// TIA Portal project "CLU" (V13) (continued)
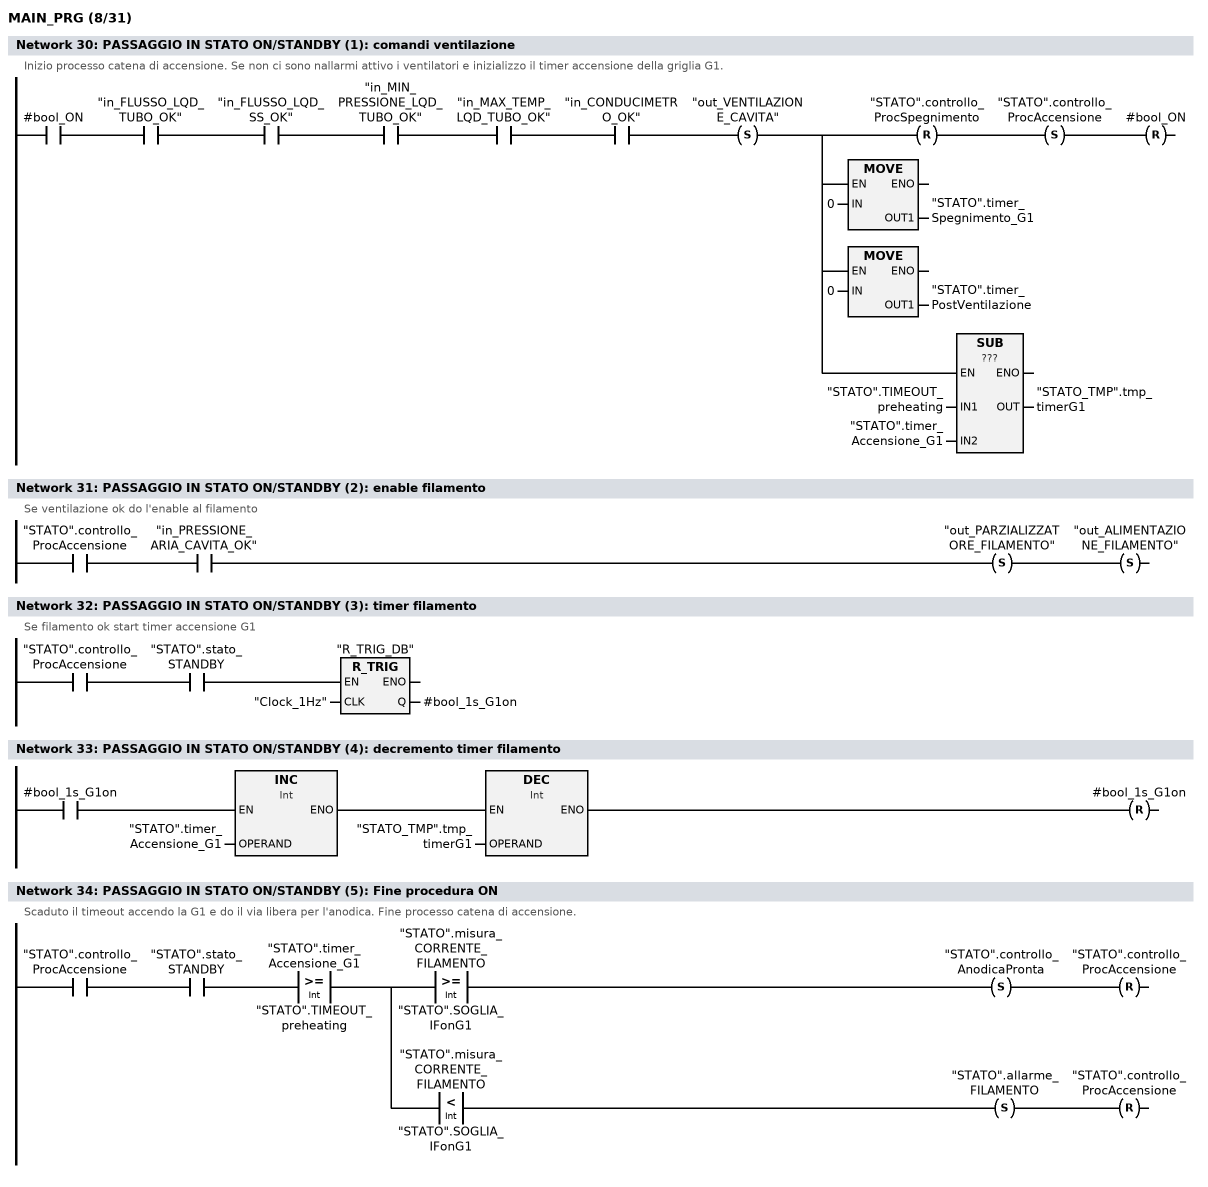
   RUNG wire#powerrail
      Contact( #bool_ON )
      Contact( "in_FLUSSO_LQD_TUBO_OK" )
      Contact( "in_FLUSSO_LQD_SS_OK" )
      Contact( "in_MIN_PRESSIONE_LQD_TUBO_OK" )
      Contact( "in_MAX_TEMP_LQD_TUBO_OK" )
      Contact( "in_CONDUCIMETRO_OK" )
      S_Coil( "out_VENTILAZIONE_CAVITA" )
      wire#w1
      R_Coil( "STATO".controllo_ProcSpegnimento )
      S_Coil( "STATO".controllo_ProcAccensione )
      R_Coil( #bool_ON )
   END_RUNG
   RUNG wire#w1
      Move(in := 0, out1 => "STATO".timer_Spegnimento_G1)
   END_RUNG
   RUNG wire#w1
      Move(in := 0, out1 => "STATO".timer_PostVentilazione)
   END_RUNG
   RUNG wire#w1
      { S7_Templates := "SrcType := ???" } Sub(in1 := "STATO".TIMEOUT_preheating, in2 := "STATO".timer_Accensione_G1, out => "STATO_TMP".tmp_timerG1)
   END_RUNG
   // the same network as SCL:
   IF #bool_ON AND "in_FLUSSO_LQD_TUBO_OK" AND "in_FLUSSO_LQD_SS_OK" AND "in_MIN_PRESSIONE_LQD_TUBO_OK" AND "in_MAX_TEMP_LQD_TUBO_OK" AND "in_CONDUCIMETRO_OK" THEN
       "out_VENTILAZIONE_CAVITA" := TRUE;
       "STATO".controllo_ProcSpegnimento := FALSE;
       "STATO".controllo_ProcAccensione := TRUE;
   END_IF;
   #_w1 := #bool_ON AND "in_FLUSSO_LQD_TUBO_OK" AND "in_FLUSSO_LQD_SS_OK" AND "in_MIN_PRESSIONE_LQD_TUBO_OK" AND "in_MAX_TEMP_LQD_TUBO_OK" AND "in_CONDUCIMETRO_OK";
   IF #_w1 THEN
       #bool_ON := FALSE;
       "STATO".timer_Spegnimento_G1 := 0;
       "STATO".timer_PostVentilazione := 0;
       "STATO_TMP".tmp_timerG1 := "STATO".TIMEOUT_preheating - "STATO".timer_Accensione_G1;
   END_IF;
END_REGION

REGION Network 31: PASSAGGIO IN STATO ON/STANDBY (2): enable filamento
   // Se ventilazione ok do l'enable al filamento
   RUNG wire#powerrail
      Contact( "STATO".controllo_ProcAccensione )
      Contact( "in_PRESSIONE_ARIA_CAVITA_OK" )
      S_Coil( "out_PARZIALIZZATORE_FILAMENTO" )
      S_Coil( "out_ALIMENTAZIONE_FILAMENTO" )
   END_RUNG
   // the same network as SCL:
   IF "STATO".controllo_ProcAccensione AND "in_PRESSIONE_ARIA_CAVITA_OK" THEN
       "out_PARZIALIZZATORE_FILAMENTO" := TRUE;
       "out_ALIMENTAZIONE_FILAMENTO" := TRUE;
   END_IF;
END_REGION

REGION Network 32: PASSAGGIO IN STATO ON/STANDBY (3): timer filamento
   // Se filamento ok start timer accensione G1
   IF "STATO".controllo_ProcAccensione AND "STATO".stato_STANDBY THEN
       "R_TRIG_DB"(CLK := "Clock_1Hz", Q => #bool_1s_G1on);   // R_TRIG
   END_IF;
END_REGION

REGION Network 33: PASSAGGIO IN STATO ON/STANDBY (4): decremento timer filamento
   RUNG wire#powerrail
      Contact( #bool_1s_G1on )
      { S7_Templates := "DestType := Int" } Inc( "STATO".timer_Accensione_G1 )
      { S7_Templates := "DestType := Int" } Dec( "STATO_TMP".tmp_timerG1 )
      R_Coil( #bool_1s_G1on )
   END_RUNG
   // the same network as SCL:
   IF #bool_1s_G1on THEN
       "STATO".timer_Accensione_G1 := "STATO".timer_Accensione_G1 + 1;
       "STATO_TMP".tmp_timerG1 := "STATO_TMP".tmp_timerG1 - 1;
       #bool_1s_G1on := FALSE;
   END_IF;
END_REGION

REGION Network 34: PASSAGGIO IN STATO ON/STANDBY (5): Fine procedura ON
   // Scaduto il timeout accendo la G1 e do il via libera per l'anodica. Fine processo catena di accensione.
   RUNG wire#powerrail
      Contact( "STATO".controllo_ProcAccensione )
      Contact( "STATO".stato_STANDBY )
      { S7_Templates := "SrcType := Int" } GE_Contact(in1 := "STATO".timer_Accensione_G1, in2 := "STATO".TIMEOUT_preheating)
      wire#w1
      { S7_Templates := "SrcType := Int" } GE_Contact(in1 := "STATO".misura_CORRENTE_FILAMENTO, in2 := "STATO".SOGLIA_IFonG1)
      S_Coil( "STATO".controllo_AnodicaPronta )
      R_Coil( "STATO".controllo_ProcAccensione )
   END_RUNG
   RUNG wire#w1
      { S7_Templates := "SrcType := Int" } LT_Contact(in1 := "STATO".misura_CORRENTE_FILAMENTO, in2 := "STATO".SOGLIA_IFonG1)
      S_Coil( "STATO".allarme_FILAMENTO )
      R_Coil( "STATO".controllo_ProcAccensione )
   END_RUNG
   // the same network as SCL:
   #_w1 := "STATO".controllo_ProcAccensione AND "STATO".stato_STANDBY AND ("STATO".timer_Accensione_G1 >= "STATO".TIMEOUT_preheating);
   IF #_w1 AND ("STATO".misura_CORRENTE_FILAMENTO >= "STATO".SOGLIA_IFonG1) THEN
       "STATO".controllo_AnodicaPronta := TRUE;
       "STATO".controllo_ProcAccensione := FALSE;
   END_IF;
   IF #_w1 AND ("STATO".misura_CORRENTE_FILAMENTO < "STATO".SOGLIA_IFonG1) THEN
       "STATO".allarme_FILAMENTO := TRUE;
       "STATO".controllo_ProcAccensione := FALSE;
   END_IF;
END_REGION

REGION Network 35: PASSAGGIO IN ANODICA ON (1): inizio accensione anodica
   // Se il processo catena di accensione è terminato posso iniziare il processo catena di accensione anodica.
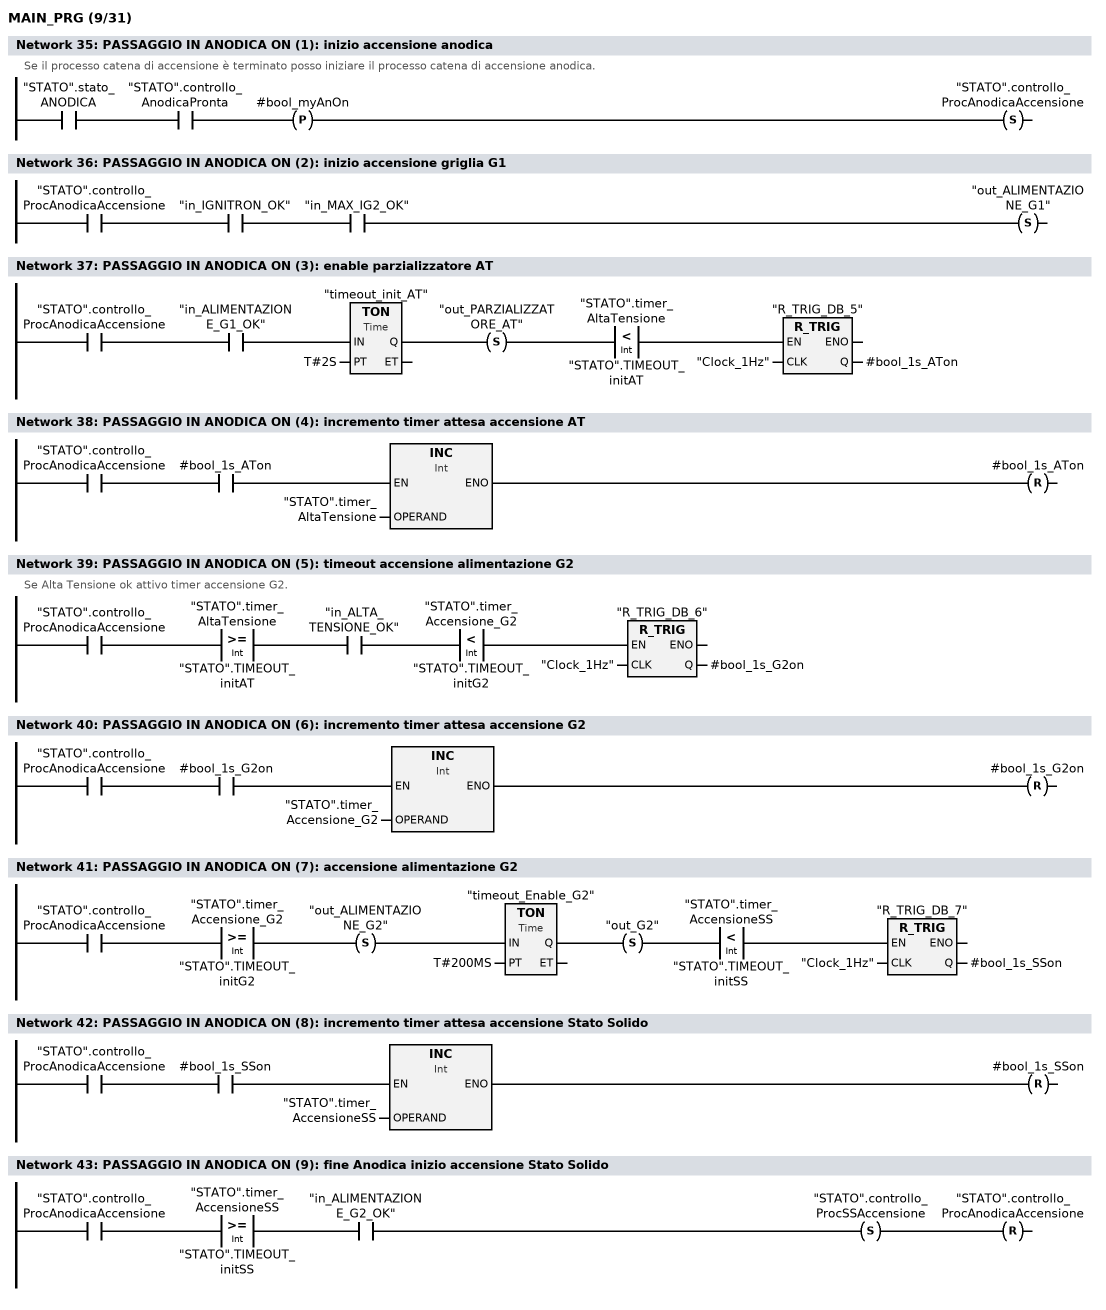
   RUNG wire#powerrail
      Contact( "STATO".stato_ANODICA )
      Contact( "STATO".controllo_AnodicaPronta )
      P_Trig( #bool_myAnOn )
      S_Coil( "STATO".controllo_ProcAnodicaAccensione )
   END_RUNG
   // the same network as SCL:
   #_w1 := "STATO".stato_ANODICA AND "STATO".controllo_AnodicaPronta;
   #_w2 := #_w1 AND NOT #bool_myAnOn;   // rising edge
   #bool_myAnOn := #_w1;
   IF #_w2 THEN "STATO".controllo_ProcAnodicaAccensione := TRUE; END_IF;
END_REGION

REGION Network 36: PASSAGGIO IN ANODICA ON (2): inizio accensione griglia G1
   RUNG wire#powerrail
      Contact( "STATO".controllo_ProcAnodicaAccensione )
      Contact( "in_IGNITRON_OK" )
      Contact( "in_MAX_IG2_OK" )
      S_Coil( "out_ALIMENTAZIONE_G1" )
   END_RUNG
   // the same network as SCL:
   IF "STATO".controllo_ProcAnodicaAccensione AND "in_IGNITRON_OK" AND "in_MAX_IG2_OK" THEN
       "out_ALIMENTAZIONE_G1" := TRUE;
   END_IF;
END_REGION

REGION Network 37: PASSAGGIO IN ANODICA ON (3): enable parzializzatore AT
   "timeout_init_AT".TON(IN := "STATO".controllo_ProcAnodicaAccensione AND "in_ALIMENTAZIONE_G1_OK", PT := T#2S);
   IF "timeout_init_AT".Q THEN "out_PARZIALIZZATORE_AT" := TRUE; END_IF;
   IF "timeout_init_AT".Q AND ("STATO".timer_AltaTensione < "STATO".TIMEOUT_initAT) THEN
       "R_TRIG_DB_5"(CLK := "Clock_1Hz", Q => #bool_1s_ATon);   // R_TRIG
   END_IF;
END_REGION

REGION Network 38: PASSAGGIO IN ANODICA ON (4): incremento timer attesa accensione AT
   RUNG wire#powerrail
      Contact( "STATO".controllo_ProcAnodicaAccensione )
      Contact( #bool_1s_ATon )
      { S7_Templates := "DestType := Int" } Inc( "STATO".timer_AltaTensione )
      R_Coil( #bool_1s_ATon )
   END_RUNG
   // the same network as SCL:
   IF "STATO".controllo_ProcAnodicaAccensione AND #bool_1s_ATon THEN
       "STATO".timer_AltaTensione := "STATO".timer_AltaTensione + 1;
       #bool_1s_ATon := FALSE;
   END_IF;
END_REGION

REGION Network 39: PASSAGGIO IN ANODICA ON (5): timeout accensione alimentazione G2
   // Se Alta Tensione ok attivo timer accensione G2.
   IF "STATO".controllo_ProcAnodicaAccensione AND ("STATO".timer_AltaTensione >= "STATO".TIMEOUT_initAT) AND "in_ALTA_TENSIONE_OK" AND ("STATO".timer_Accensione_G2 < "STATO".TIMEOUT_initG2) THEN
       "R_TRIG_DB_6"(CLK := "Clock_1Hz", Q => #bool_1s_G2on);   // R_TRIG
   END_IF;
END_REGION

REGION Network 40: PASSAGGIO IN ANODICA ON (6): incremento timer attesa accensione G2
   RUNG wire#powerrail
      Contact( "STATO".controllo_ProcAnodicaAccensione )
      Contact( #bool_1s_G2on )
      { S7_Templates := "DestType := Int" } Inc( "STATO".timer_Accensione_G2 )
      R_Coil( #bool_1s_G2on )
   END_RUNG
   // the same network as SCL:
   IF "STATO".controllo_ProcAnodicaAccensione AND #bool_1s_G2on THEN
       "STATO".timer_Accensione_G2 := "STATO".timer_Accensione_G2 + 1;
       #bool_1s_G2on := FALSE;
   END_IF;
END_REGION

REGION Network 41: PASSAGGIO IN ANODICA ON (7): accensione alimentazione G2
   #_w1 := "STATO".controllo_ProcAnodicaAccensione AND ("STATO".timer_Accensione_G2 >= "STATO".TIMEOUT_initG2);
   IF #_w1 THEN "out_ALIMENTAZIONE_G2" := TRUE; END_IF;
   "timeout_Enable_G2".TON(IN := #_w1, PT := T#200MS);
   IF "timeout_Enable_G2".Q THEN "out_G2" := TRUE; END_IF;
   IF "timeout_Enable_G2".Q AND ("STATO".timer_AccensioneSS < "STATO".TIMEOUT_initSS) THEN
       "R_TRIG_DB_7"(CLK := "Clock_1Hz", Q => #bool_1s_SSon);   // R_TRIG
   END_IF;
END_REGION

REGION Network 42: PASSAGGIO IN ANODICA ON (8): incremento timer attesa accensione Stato Solido
   RUNG wire#powerrail
      Contact( "STATO".controllo_ProcAnodicaAccensione )
      Contact( #bool_1s_SSon )
      { S7_Templates := "DestType := Int" } Inc( "STATO".timer_AccensioneSS )
      R_Coil( #bool_1s_SSon )
   END_RUNG
   // the same network as SCL:
   IF "STATO".controllo_ProcAnodicaAccensione AND #bool_1s_SSon THEN
       "STATO".timer_AccensioneSS := "STATO".timer_AccensioneSS + 1;
       #bool_1s_SSon := FALSE;
   END_IF;
END_REGION

REGION Network 43: PASSAGGIO IN ANODICA ON (9): fine Anodica inizio accensione Stato Solido
   RUNG wire#powerrail
      Contact( "STATO".controllo_ProcAnodicaAccensione )
      { S7_Templates := "SrcType := Int" } GE_Contact(in1 := "STATO".timer_AccensioneSS, in2 := "STATO".TIMEOUT_initSS)
      Contact( "in_ALIMENTAZIONE_G2_OK" )
      S_Coil( "STATO".controllo_ProcSSAccensione )
      R_Coil( "STATO".controllo_ProcAnodicaAccensione )
   END_RUNG
   // the same network as SCL:
   IF "STATO".controllo_ProcAnodicaAccensione AND ("STATO".timer_AccensioneSS >= "STATO".TIMEOUT_initSS) AND "in_ALIMENTAZIONE_G2_OK" THEN
       "STATO".controllo_ProcSSAccensione := TRUE;
       "STATO".controllo_ProcAnodicaAccensione := FALSE;
   END_IF;
END_REGION

REGION Network 44: ACCENSIONE STATO SOLIDO (1): accensione amplificatore (impulsivo) AMP 1
   // Se modalità  impulsiva attiva accendo gli amplificatori e attivo timer accensione driver.
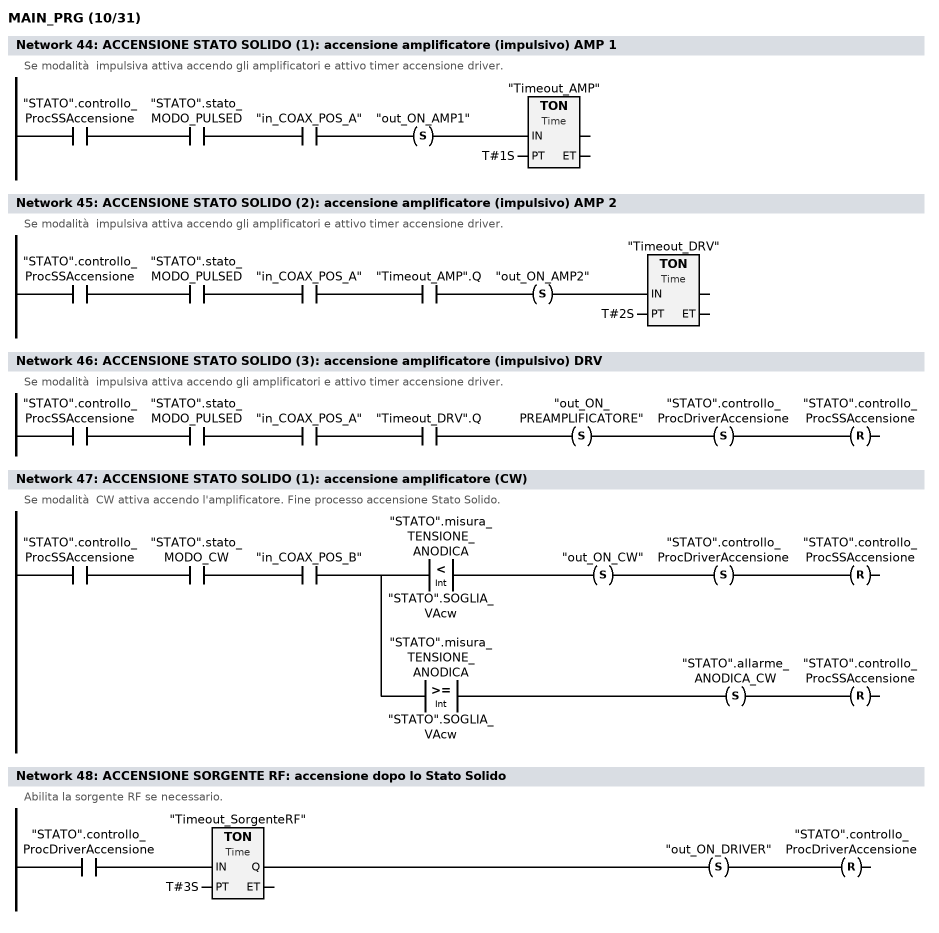
   #_w1 := "STATO".controllo_ProcSSAccensione AND "STATO".stato_MODO_PULSED AND "in_COAX_POS_A";
   IF #_w1 THEN "out_ON_AMP1" := TRUE; END_IF;
   "Timeout_AMP".TON(IN := #_w1, PT := T#1S);
END_REGION

REGION Network 45: ACCENSIONE STATO SOLIDO (2): accensione amplificatore (impulsivo) AMP 2
   // Se modalità  impulsiva attiva accendo gli amplificatori e attivo timer accensione driver.
   #_w1 := "STATO".controllo_ProcSSAccensione AND "STATO".stato_MODO_PULSED AND "in_COAX_POS_A" AND "Timeout_AMP".Q;
   IF #_w1 THEN "out_ON_AMP2" := TRUE; END_IF;
   "Timeout_DRV".TON(IN := #_w1, PT := T#2S);
END_REGION

REGION Network 46: ACCENSIONE STATO SOLIDO (3): accensione amplificatore (impulsivo) DRV
   // Se modalità  impulsiva attiva accendo gli amplificatori e attivo timer accensione driver.
   RUNG wire#powerrail
      Contact( "STATO".controllo_ProcSSAccensione )
      Contact( "STATO".stato_MODO_PULSED )
      Contact( "in_COAX_POS_A" )
      Contact( "Timeout_DRV".Q )
      S_Coil( "out_ON_PREAMPLIFICATORE" )
      S_Coil( "STATO".controllo_ProcDriverAccensione )
      R_Coil( "STATO".controllo_ProcSSAccensione )
   END_RUNG
   // the same network as SCL:
   IF "STATO".controllo_ProcSSAccensione AND "STATO".stato_MODO_PULSED AND "in_COAX_POS_A" AND "Timeout_DRV".Q THEN
       "out_ON_PREAMPLIFICATORE" := TRUE;
       "STATO".controllo_ProcDriverAccensione := TRUE;
       "STATO".controllo_ProcSSAccensione := FALSE;
   END_IF;
END_REGION

REGION Network 47: ACCENSIONE STATO SOLIDO (1): accensione amplificatore (CW)
   // Se modalità  CW attiva accendo l'amplificatore. Fine processo accensione Stato Solido.
   RUNG wire#powerrail
      Contact( "STATO".controllo_ProcSSAccensione )
      Contact( "STATO".stato_MODO_CW )
      Contact( "in_COAX_POS_B" )
      wire#w1
      { S7_Templates := "SrcType := Int" } LT_Contact(in1 := "STATO".misura_TENSIONE_ANODICA, in2 := "STATO".SOGLIA_VAcw)
      S_Coil( "out_ON_CW" )
      S_Coil( "STATO".controllo_ProcDriverAccensione )
      R_Coil( "STATO".controllo_ProcSSAccensione )
   END_RUNG
   RUNG wire#w1
      { S7_Templates := "SrcType := Int" } GE_Contact(in1 := "STATO".misura_TENSIONE_ANODICA, in2 := "STATO".SOGLIA_VAcw)
      S_Coil( "STATO".allarme_ANODICA_CW )
      R_Coil( "STATO".controllo_ProcSSAccensione )
   END_RUNG
   // the same network as SCL:
   #_w1 := "STATO".controllo_ProcSSAccensione AND "STATO".stato_MODO_CW AND "in_COAX_POS_B";
   IF #_w1 AND ("STATO".misura_TENSIONE_ANODICA < "STATO".SOGLIA_VAcw) THEN
       "out_ON_CW" := TRUE;
       "STATO".controllo_ProcDriverAccensione := TRUE;
       "STATO".controllo_ProcSSAccensione := FALSE;
   END_IF;
   IF #_w1 AND ("STATO".misura_TENSIONE_ANODICA >= "STATO".SOGLIA_VAcw) THEN
       "STATO".allarme_ANODICA_CW := TRUE;
       "STATO".controllo_ProcSSAccensione := FALSE;
   END_IF;
END_REGION

REGION Network 48: ACCENSIONE SORGENTE RF: accensione dopo lo Stato Solido
   // Abilita la sorgente RF se necessario.
   "Timeout_SorgenteRF".TON(IN := "STATO".controllo_ProcDriverAccensione, PT := T#3S);
   IF "Timeout_SorgenteRF".Q THEN
       "out_ON_DRIVER" := TRUE;
       "STATO".controllo_ProcDriverAccensione := FALSE;
   END_IF;
END_REGION

REGION Network 49: PASSAGGIO IN ANODICA OFF (1): spegnimento Stato Solido e alimentazione G2
   // Spengo Stato Solido (CW o impulsivo) e alimentazione G2. Inizio processo catena di spegnimento Anodica.
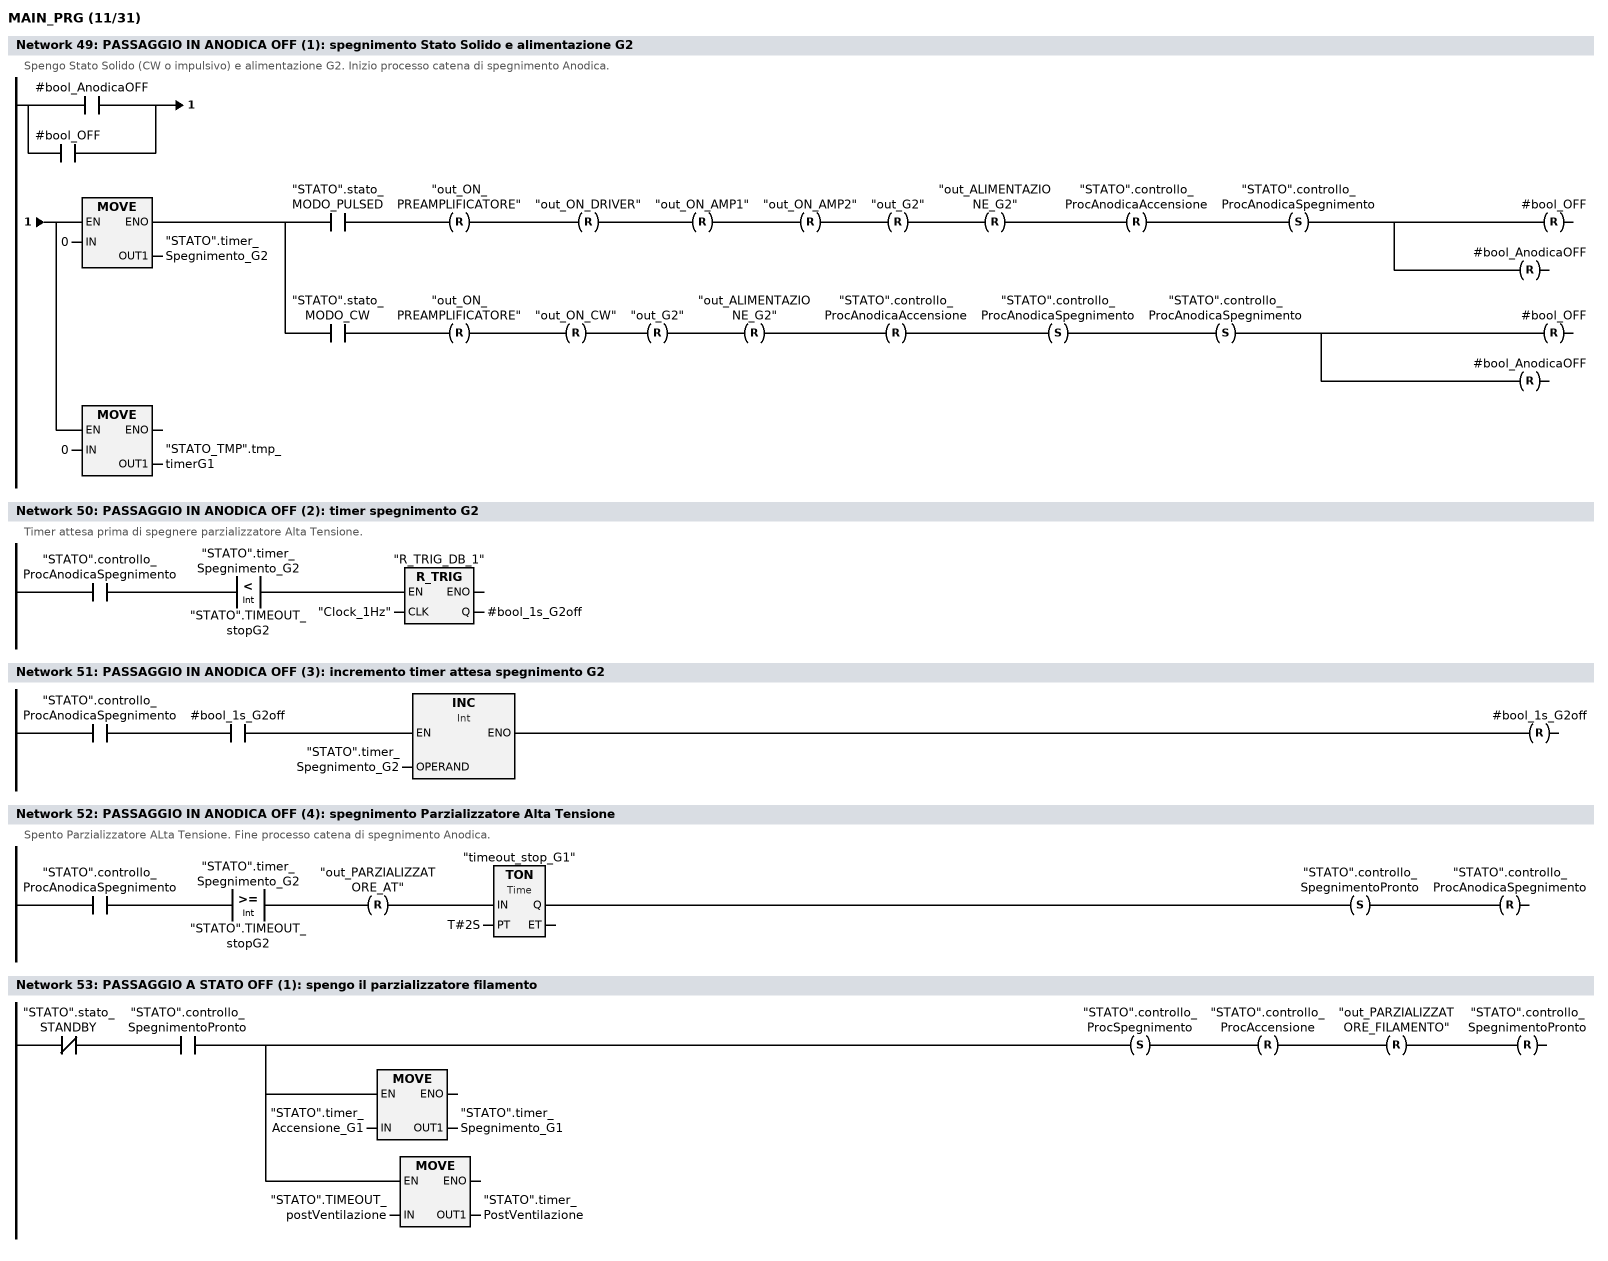
   RUNG wire#powerrail
      Contact( #bool_AnodicaOFF )
      wire#w1
      Move(in := 0, out1 => "STATO".timer_Spegnimento_G2)
      wire#w2
      Contact( "STATO".stato_MODO_PULSED )
      R_Coil( "out_ON_PREAMPLIFICATORE" )
      R_Coil( "out_ON_DRIVER" )
      R_Coil( "out_ON_AMP1" )
      R_Coil( "out_ON_AMP2" )
      R_Coil( "out_G2" )
      R_Coil( "out_ALIMENTAZIONE_G2" )
      R_Coil( "STATO".controllo_ProcAnodicaAccensione )
      S_Coil( "STATO".controllo_ProcAnodicaSpegnimento )
      wire#w3
      R_Coil( #bool_OFF )
   END_RUNG
   RUNG wire#powerrail
      Contact( #bool_OFF )
   END_RUNG wire#w1
   RUNG wire#w3
      R_Coil( #bool_AnodicaOFF )
   END_RUNG
   RUNG wire#w2
      Contact( "STATO".stato_MODO_CW )
      R_Coil( "out_ON_PREAMPLIFICATORE" )
      R_Coil( "out_ON_CW" )
      R_Coil( "out_G2" )
      R_Coil( "out_ALIMENTAZIONE_G2" )
      R_Coil( "STATO".controllo_ProcAnodicaAccensione )
      S_Coil( "STATO".controllo_ProcAnodicaSpegnimento )
      S_Coil( "STATO".controllo_ProcAnodicaSpegnimento )
      wire#w4
      R_Coil( #bool_OFF )
   END_RUNG
   RUNG wire#w4
      R_Coil( #bool_AnodicaOFF )
   END_RUNG
   RUNG wire#w1
      Move(in := 0, out1 => "STATO_TMP".tmp_timerG1)
   END_RUNG
   // the same network as SCL:
   #_w1 := #bool_AnodicaOFF OR #bool_OFF;
   IF #_w1 THEN "STATO".timer_Spegnimento_G2 := 0; END_IF;
   IF #_w1 AND "STATO".stato_MODO_PULSED THEN
       "out_ON_PREAMPLIFICATORE" := FALSE;
       "out_ON_DRIVER" := FALSE;
       "out_ON_AMP1" := FALSE;
       "out_ON_AMP2" := FALSE;
       "out_G2" := FALSE;
       "out_ALIMENTAZIONE_G2" := FALSE;
       "STATO".controllo_ProcAnodicaAccensione := FALSE;
       "STATO".controllo_ProcAnodicaSpegnimento := TRUE;
       #bool_OFF := FALSE;
       #bool_AnodicaOFF := FALSE;
   END_IF;
   IF #_w1 AND "STATO".stato_MODO_CW THEN
       "out_ON_PREAMPLIFICATORE" := FALSE;
       "out_ON_CW" := FALSE;
       "out_G2" := FALSE;
       "out_ALIMENTAZIONE_G2" := FALSE;
       "STATO".controllo_ProcAnodicaAccensione := FALSE;
       "STATO".controllo_ProcAnodicaSpegnimento := TRUE;
       "STATO".controllo_ProcAnodicaSpegnimento := TRUE;
       #bool_OFF := FALSE;
       #bool_AnodicaOFF := FALSE;
   END_IF;
   IF #_w1 THEN "STATO_TMP".tmp_timerG1 := 0; END_IF;
END_REGION

REGION Network 50: PASSAGGIO IN ANODICA OFF (2): timer spegnimento G2
   // Timer attesa prima di spegnere parzializzatore Alta Tensione.
   IF "STATO".controllo_ProcAnodicaSpegnimento AND ("STATO".timer_Spegnimento_G2 < "STATO".TIMEOUT_stopG2) THEN
       "R_TRIG_DB_1"(CLK := "Clock_1Hz", Q => #bool_1s_G2off);   // R_TRIG
   END_IF;
END_REGION

REGION Network 51: PASSAGGIO IN ANODICA OFF (3): incremento timer attesa spegnimento G2
   RUNG wire#powerrail
      Contact( "STATO".controllo_ProcAnodicaSpegnimento )
      Contact( #bool_1s_G2off )
      { S7_Templates := "DestType := Int" } Inc( "STATO".timer_Spegnimento_G2 )
      R_Coil( #bool_1s_G2off )
   END_RUNG
   // the same network as SCL:
   IF "STATO".controllo_ProcAnodicaSpegnimento AND #bool_1s_G2off THEN
       "STATO".timer_Spegnimento_G2 := "STATO".timer_Spegnimento_G2 + 1;
       #bool_1s_G2off := FALSE;
   END_IF;
END_REGION

REGION Network 52: PASSAGGIO IN ANODICA OFF (4): spegnimento Parzializzatore Alta Tensione
   // Spento Parzializzatore ALta Tensione. Fine processo catena di spegnimento Anodica.
   #_w1 := "STATO".controllo_ProcAnodicaSpegnimento AND ("STATO".timer_Spegnimento_G2 >= "STATO".TIMEOUT_stopG2);
   IF #_w1 THEN "out_PARZIALIZZATORE_AT" := FALSE; END_IF;
   "timeout_stop_G1".TON(IN := #_w1, PT := T#2S);
   IF "timeout_stop_G1".Q THEN
       "STATO".controllo_SpegnimentoPronto := TRUE;
       "STATO".controllo_ProcAnodicaSpegnimento := FALSE;
   END_IF;
END_REGION

REGION Network 53: PASSAGGIO A STATO OFF (1): spengo il parzializzatore filamento
   RUNG wire#powerrail
      I_Contact( "STATO".stato_STANDBY )
      Contact( "STATO".controllo_SpegnimentoPronto )
      wire#w1
      S_Coil( "STATO".controllo_ProcSpegnimento )
      R_Coil( "STATO".controllo_ProcAccensione )
      R_Coil( "out_PARZIALIZZATORE_FILAMENTO" )
      R_Coil( "STATO".controllo_SpegnimentoPronto )
   END_RUNG
   RUNG wire#w1
      Move(in := "STATO".timer_Accensione_G1, out1 => "STATO".timer_Spegnimento_G1)
   END_RUNG
   RUNG wire#w1
      Move(in := "STATO".TIMEOUT_postVentilazione, out1 => "STATO".timer_PostVentilazione)
   END_RUNG
   // the same network as SCL:
   IF NOT "STATO".stato_STANDBY AND "STATO".controllo_SpegnimentoPronto THEN
       "STATO".controllo_ProcSpegnimento := TRUE;
       "STATO".controllo_ProcAccensione := FALSE;
       "out_PARZIALIZZATORE_FILAMENTO" := FALSE;
   END_IF;
   #_w1 := NOT "STATO".stato_STANDBY AND "STATO".controllo_SpegnimentoPronto;
   IF #_w1 THEN
       "STATO".controllo_SpegnimentoPronto := FALSE;
       "STATO".timer_Spegnimento_G1 := "STATO".timer_Accensione_G1;
       "STATO".timer_PostVentilazione := "STATO".TIMEOUT_postVentilazione;
   END_IF;
END_REGION

REGION Network 54: PASSAGGIO A STATO OFF (2): attesa spegnimento alimentazione Filamento
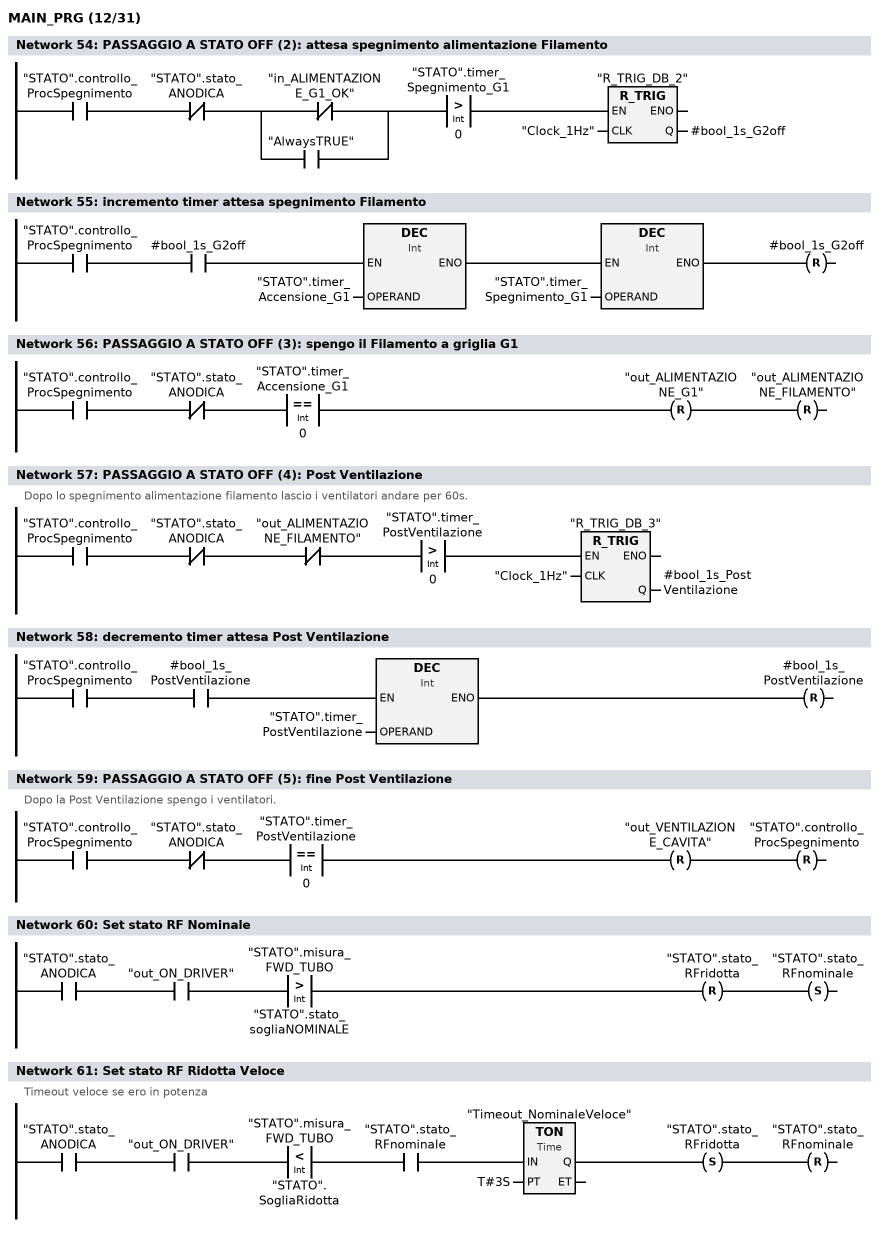
   IF "STATO".controllo_ProcSpegnimento AND NOT "STATO".stato_ANODICA AND (NOT "in_ALIMENTAZIONE_G1_OK" OR "AlwaysTRUE") AND ("STATO".timer_Spegnimento_G1 > 0) THEN
       "R_TRIG_DB_2"(CLK := "Clock_1Hz", Q => #bool_1s_G2off);   // R_TRIG
   END_IF;
END_REGION

REGION Network 55: incremento timer attesa spegnimento Filamento
   RUNG wire#powerrail
      Contact( "STATO".controllo_ProcSpegnimento )
      Contact( #bool_1s_G2off )
      { S7_Templates := "DestType := Int" } Dec( "STATO".timer_Accensione_G1 )
      { S7_Templates := "DestType := Int" } Dec( "STATO".timer_Spegnimento_G1 )
      R_Coil( #bool_1s_G2off )
   END_RUNG
   // the same network as SCL:
   IF "STATO".controllo_ProcSpegnimento AND #bool_1s_G2off THEN
       "STATO".timer_Accensione_G1 := "STATO".timer_Accensione_G1 - 1;
       "STATO".timer_Spegnimento_G1 := "STATO".timer_Spegnimento_G1 - 1;
       #bool_1s_G2off := FALSE;
   END_IF;
END_REGION

REGION Network 56: PASSAGGIO A STATO OFF (3): spengo il Filamento a griglia G1
   RUNG wire#powerrail
      Contact( "STATO".controllo_ProcSpegnimento )
      I_Contact( "STATO".stato_ANODICA )
      { S7_Templates := "SrcType := Int" } EQ_Contact(in1 := "STATO".timer_Accensione_G1, in2 := 0)
      R_Coil( "out_ALIMENTAZIONE_G1" )
      R_Coil( "out_ALIMENTAZIONE_FILAMENTO" )
   END_RUNG
   // the same network as SCL:
   IF "STATO".controllo_ProcSpegnimento AND NOT "STATO".stato_ANODICA AND ("STATO".timer_Accensione_G1 = 0) THEN
       "out_ALIMENTAZIONE_G1" := FALSE;
       "out_ALIMENTAZIONE_FILAMENTO" := FALSE;
   END_IF;
END_REGION

REGION Network 57: PASSAGGIO A STATO OFF (4): Post Ventilazione
   // Dopo lo spegnimento alimentazione filamento lascio i ventilatori andare per 60s.
   IF "STATO".controllo_ProcSpegnimento AND NOT "STATO".stato_ANODICA AND NOT "out_ALIMENTAZIONE_FILAMENTO" AND ("STATO".timer_PostVentilazione > 0) THEN
       "R_TRIG_DB_3"(CLK := "Clock_1Hz", Q => #bool_1s_PostVentilazione);   // R_TRIG
   END_IF;
END_REGION

REGION Network 58: decremento timer attesa Post Ventilazione
   RUNG wire#powerrail
      Contact( "STATO".controllo_ProcSpegnimento )
      Contact( #bool_1s_PostVentilazione )
      { S7_Templates := "DestType := Int" } Dec( "STATO".timer_PostVentilazione )
      R_Coil( #bool_1s_PostVentilazione )
   END_RUNG
   // the same network as SCL:
   IF "STATO".controllo_ProcSpegnimento AND #bool_1s_PostVentilazione THEN
       "STATO".timer_PostVentilazione := "STATO".timer_PostVentilazione - 1;
       #bool_1s_PostVentilazione := FALSE;
   END_IF;
END_REGION

REGION Network 59: PASSAGGIO A STATO OFF (5): fine Post Ventilazione
   // Dopo la Post Ventilazione spengo i ventilatori.
   RUNG wire#powerrail
      Contact( "STATO".controllo_ProcSpegnimento )
      I_Contact( "STATO".stato_ANODICA )
      { S7_Templates := "SrcType := Int" } EQ_Contact(in1 := "STATO".timer_PostVentilazione, in2 := 0)
      R_Coil( "out_VENTILAZIONE_CAVITA" )
      R_Coil( "STATO".controllo_ProcSpegnimento )
   END_RUNG
   // the same network as SCL:
   IF "STATO".controllo_ProcSpegnimento AND NOT "STATO".stato_ANODICA AND ("STATO".timer_PostVentilazione = 0) THEN
       "out_VENTILAZIONE_CAVITA" := FALSE;
       "STATO".controllo_ProcSpegnimento := FALSE;
   END_IF;
END_REGION

REGION Network 60: Set stato RF Nominale
   RUNG wire#powerrail
      Contact( "STATO".stato_ANODICA )
      Contact( "out_ON_DRIVER" )
      { S7_Templates := "SrcType := Int" } GT_Contact(in1 := "STATO".misura_FWD_TUBO, in2 := "STATO".stato_sogliaNOMINALE)
      R_Coil( "STATO".stato_RFridotta )
      S_Coil( "STATO".stato_RFnominale )
   END_RUNG
   // the same network as SCL:
   IF "STATO".stato_ANODICA AND "out_ON_DRIVER" AND ("STATO".misura_FWD_TUBO > "STATO".stato_sogliaNOMINALE) THEN
       "STATO".stato_RFridotta := FALSE;
       "STATO".stato_RFnominale := TRUE;
   END_IF;
END_REGION

REGION Network 61: Set stato RF Ridotta Veloce
   // Timeout veloce se ero in potenza
   "Timeout_NominaleVeloce".TON(IN := "STATO".stato_ANODICA AND "out_ON_DRIVER" AND ("STATO".misura_FWD_TUBO < "STATO".SogliaRidotta) AND "STATO".stato_RFnominale,
                           PT := T#3S);
   IF "Timeout_NominaleVeloce".Q THEN
       "STATO".stato_RFridotta := TRUE;
       "STATO".stato_RFnominale := FALSE;
   END_IF;
END_REGION

REGION Network 62: Set stato RF Ridotta
   // Timeout lento se non ero in potenza